// TIA Portal project "Log Control" (V20)

(* hardware
DEVICE "S7-1500/ET200MP station_1"  S7-1500 station
   slot 0: "Rail_0"  Rack  6ES7 590-1***0-0AA0
   slot 1: "PLC_1"  CPU 1518T-3 PN  6ES7 518-3TT10-0AB0  V4.0
      slot 3: "CPU display_1"  6ES7591-1BA00-0AA0
      slot 32768: "PROFINET interface_1"  X1
         slot 32769: "Port_1"  X1 P1
         slot 32770: "Port_2"  X1 P2
      slot 33024: "PROFINET interface_2"  X2
         slot 33025: "Port_1"  X2 P1
         slot 33026: "Port_2"  X2 P2
      slot 33280: "PROFINET interface GBIT_3"  X3
         slot 33281: "Port_1"  X3 P1
      slot 34817: "Virtual CP interface port_1"  Virtual CP interface port  Virtual CP interface port FW V4.0
DEVICE "LogHMI"  KTP700 Basic PN
   slot 0: "anit-hmi"  KTP700 Basic PN  6AV2 123-2GB03-0AX0  17.0.0.0
   slot 1: "HMI_RT_1"  KTP700 Basic PN  6AV2 123-2GB03-0AX0  17.0.0.0
   slot 5: "anit-hmi.IE_CP_1"  PROFINET Interface  17.0.0.0
      slot 1: "PROFINET Interface_1"  PROFINET Interface
         slot 1: "Port_1"  Port
*)

// ===== PLC "PLC_1"  CPU 1518T-3 PN =====
// protected blocks, not shown: "Log Control FC"

VAR_GLOBAL   // PLC tag table "Default tag table"
   "Tag_1" AT %M45.0 : Bool;
   "Tag_2" AT %M0.0 : Bool;
   "Tag_3" AT %M0.1 : Bool;
   "Tag_4" AT %M47.0 : Bool;
   "Tag_5" AT %M31.0 : Bool;
END_VAR

TYPE "LogControlUDT"
   STRUCT
      Settings : Struct
         "In Min" : Int := 0;
         "In Max" : Int := 100;
         "Out Min" : Real := 0.0;
         "Out Max" : Real := 100.0;
         "Log Repeat time" : Time := T#1s;
      END_STRUCT;
      "Worning Control" : Array[1..10] of Struct
         Text : String[20];
         MinValue : Real;
         MaxValue : Real;
      END_STRUCT;
      "Prescription Control" : Struct
         "Aktif Reçete" : Struct
            "Tarih/Saat" : DTL;
            Value : Real;
            Text : String;
         END_STRUCT;
         "Reçete Göstege" : Struct
            No : Array[0..10] of Int;
            "Tarih/Saat" : Array[0..10] of DTL;
            Value : Array[0..10] of Real;
            Text : Array[0..10] of String;
         END_STRUCT;
         T_ADD_Out : DTL;
         RET_Val_Out : DTL;
         p : Bool;
         "OP No" : Int;
         "OP Artı" : Bool;
         "OP Eksi" : Bool;
         "Gösterge No" : Int;
         "Gösterge Artı" : Bool;
         "Gösterge Eksi" : Bool;
         Log_Wride : Bool;
      END_STRUCT;
      Prescription : Array[0..101] of Struct
         "Tarih/Saat" : DTL;
         Value : Real;
         Text : String;
      END_STRUCT;
   END_STRUCT;
   // "Worning Control"[1].MinValue := 0.0;
   // "Worning Control"[1].MaxValue := 10.0;
   // "Worning Control"[1].Text := 'Value1';
   // "Worning Control"[2].Text := 'Value2';
   // "Worning Control"[2].MinValue := 10.0;
   // "Worning Control"[2].MaxValue := 20.0;
   // "Worning Control"[3].Text := 'Value3';
   // "Worning Control"[3].MinValue := 20.0;
   // "Worning Control"[3].MaxValue := 30.0;
   // "Worning Control"[4].Text := 'Value4';
   // "Worning Control"[4].MinValue := 30.0;
   // "Worning Control"[4].MaxValue := 40.0;
   // "Worning Control"[5].Text := 'Value5';
   // "Worning Control"[5].MinValue := 40.0;
   // "Worning Control"[5].MaxValue := 50.0;
   // "Worning Control"[6].Text := 'Value6';
   // "Worning Control"[6].MinValue := 50.0;
   // "Worning Control"[6].MaxValue := 60.0;
   // "Worning Control"[7].Text := 'Value7';
   // "Worning Control"[7].MinValue := 60.0;
   // "Worning Control"[7].MaxValue := 70.0;
   // "Worning Control"[8].Text := 'Value8';
   // "Worning Control"[8].MinValue := 70.0;
   // "Worning Control"[8].MaxValue := 80.0;
   // "Worning Control"[9].Text := 'Value9';
   // "Worning Control"[9].MinValue := 80.0;
   // "Worning Control"[9].MaxValue := 90.0;
   // "Worning Control"[10].Text := 'Value10';
   // "Worning Control"[10].MinValue := 90.0;
   // "Worning Control"[10].MaxValue := 100.0;
END_TYPE

DATA_BLOCK "Log Control DB"   // DB1
{ S7_Optimized_Access := 'TRUE' }
VERSION : 0.1
   VAR
      LogData : "LogControlUDT";
   END_VAR
BEGIN
END_DATA_BLOCK

// folder: 99-FuncLibrary

DATA_BLOCK "Value_1"   // DB4
{ S7_Optimized_Access := 'TRUE' }
VERSION : 0.1
   VAR
      InValue : Int;
      OutValue : Int;
      OutTime : DTL;
      OutText : String;
   END_VAR
BEGIN
END_DATA_BLOCK

// folder: System blocks/Program resources

DATA_BLOCK "IEC_Timer_0_DB"   // DB2
{ S7_Optimized_Access := 'TRUE' }
AUTHOR : Simatic
FAMILY : IEC
NAME : IEC_TMR
VERSION : 1.0
// stored: InstanceOfName IEC_TIMER
"IEC_TIMER"
BEGIN
END_DATA_BLOCK

DATA_BLOCK "IEC_Counter_0_DB"   // DB3
{ S7_Optimized_Access := 'TRUE' }
AUTHOR : Simatic
FAMILY : IEC
NAME : CNTR
VERSION : 1.0
// stored: InstanceOfName IEC_COUNTER
"IEC_COUNTER"
BEGIN
END_DATA_BLOCK

DATA_BLOCK "Value"   // DB5
{ S7_Optimized_Access := 'TRUE' }
AUTHOR : Simatic
FAMILY : IEC
NAME : IEC_TMR
VERSION : 1.0
// stored: InstanceOfName IEC_TIMER
"IEC_TIMER"
BEGIN
END_DATA_BLOCK

// folder: (top level)

ORGANIZATION_BLOCK "Main"   // OB1, LAD, ProgramCycle
TITLE = "Main Program Sweep (Cycle)"
{ S7_Optimized_Access := 'TRUE' }
VERSION : 0.1
   VAR_INPUT
      Initial_Call : Bool;   // Initial call of this OB
      Remanence : Bool;   // =True, if remanent data are available
   END_VAR
   VAR_TEMP
      Reset : Bool;
   END_VAR
   VAR_TEMP   // added for the SCL form of the ladder/FBD networks
      _w1 : Bool;
   END_VAR
BEGIN

REGION Network 1
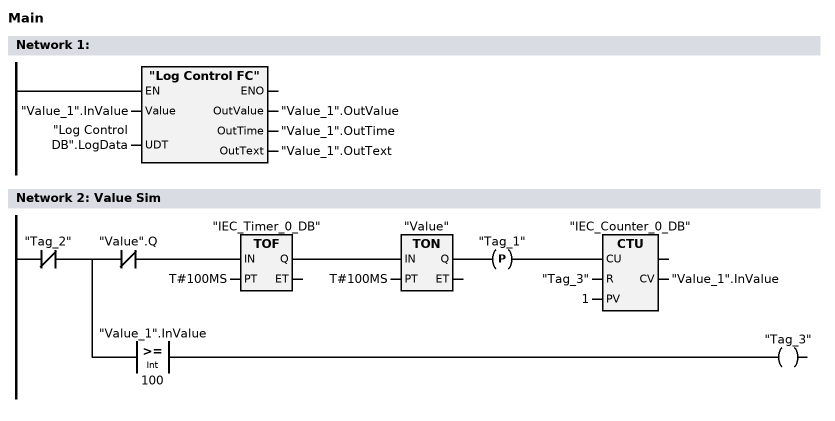
   RUNG wire#powerrail
      "Log Control FC"(Value := "Value_1".InValue, UDT := "Log Control DB".LogData, OutValue => "Value_1".OutValue, OutTime => "Value_1".OutTime, OutText => "Value_1".OutText)
   END_RUNG
   // the same network as SCL:
   "Log Control FC"(Value := "Value_1".InValue,
                    UDT := "Log Control DB".LogData,
                    OutValue => "Value_1".OutValue,
                    OutTime => "Value_1".OutTime,
                    OutText => "Value_1".OutText);
END_REGION

REGION Network 2: Value Sim
   "IEC_Timer_0_DB".TOF(IN := NOT "Tag_2" AND NOT "Value".Q, PT := T#100MS);
   "Value".TON(IN := "IEC_Timer_0_DB".Q, PT := T#100MS);
   #_w1 := "Value".Q AND NOT "Tag_1";   // rising edge
   "Tag_1" := "Value".Q;
   "IEC_Counter_0_DB".CTU(CU := #_w1, R := "Tag_3", PV := 1, CV => "Value_1".InValue);
   "Tag_3" := NOT "Tag_2" AND ("Value_1".InValue >= 100);
END_REGION
END_ORGANIZATION_BLOCK

(* ===== HMI "HMI_RT_1" =====
system functions are stored by id; their names below are inferred from use
connection "HMI_Connection_1": ETHERNET, SMART_S7_1500_OMS

HMI tags "Default tag table"
   "Log Control DB_LogData_Prescription Control_Reçete Göstege_No{1}" : Int = PLC "Log Control DB".LogData."Prescription Control"."Reçete Göstege".No[1], 100 ms
   "Log Control DB_LogData_Prescription Control_Reçete Göstege_No{2}" : Int = PLC "Log Control DB".LogData."Prescription Control"."Reçete Göstege".No[2], 100 ms
   "Log Control DB_LogData_Prescription Control_Reçete Göstege_No{3}" : Int = PLC "Log Control DB".LogData."Prescription Control"."Reçete Göstege".No[3], 100 ms
   "Log Control DB_LogData_Prescription Control_Reçete Göstege_No{4}" : Int = PLC "Log Control DB".LogData."Prescription Control"."Reçete Göstege".No[4], 100 ms
   "Log Control DB_LogData_Prescription Control_Reçete Göstege_No{5}" : Int = PLC "Log Control DB".LogData."Prescription Control"."Reçete Göstege".No[5], 100 ms
   "Log Control DB_LogData_Prescription Control_Reçete Göstege_No{6}" : Int = PLC "Log Control DB".LogData."Prescription Control"."Reçete Göstege".No[6], 100 ms
   "Log Control DB_LogData_Prescription Control_Reçete Göstege_No{7}" : Int = PLC "Log Control DB".LogData."Prescription Control"."Reçete Göstege".No[7], 100 ms
   "Log Control DB_LogData_Prescription Control_Reçete Göstege_No{8}" : Int = PLC "Log Control DB".LogData."Prescription Control"."Reçete Göstege".No[8], 100 ms
   "Log Control DB_LogData_Prescription Control_Reçete Göstege_No{9}" : Int = PLC "Log Control DB".LogData."Prescription Control"."Reçete Göstege".No[9], 100 ms
   "Log Control DB_LogData_Prescription Control_Reçete Göstege_No{10}" : Int = PLC "Log Control DB".LogData."Prescription Control"."Reçete Göstege".No[10], 100 ms
   "Log Control DB_LogData_Prescription Control_Reçete Göstege_Tarih/Saat{1}" : DTL = PLC "Log Control DB".LogData."Prescription Control"."Reçete Göstege".Tarih/Saat[1], 100 ms
   "Log Control DB_LogData_Prescription Control_Reçete Göstege_Tarih/Saat{2}" : DTL = PLC "Log Control DB".LogData."Prescription Control"."Reçete Göstege".Tarih/Saat[2], 100 ms
   "Log Control DB_LogData_Prescription Control_Reçete Göstege_Tarih/Saat{3}" : DTL = PLC "Log Control DB".LogData."Prescription Control"."Reçete Göstege".Tarih/Saat[3], 100 ms
   "Log Control DB_LogData_Prescription Control_Reçete Göstege_Tarih/Saat{4}" : DTL = PLC "Log Control DB".LogData."Prescription Control"."Reçete Göstege".Tarih/Saat[4], 100 ms
   "Log Control DB_LogData_Prescription Control_Reçete Göstege_Tarih/Saat{5}" : DTL = PLC "Log Control DB".LogData."Prescription Control"."Reçete Göstege".Tarih/Saat[5], 100 ms
   "Log Control DB_LogData_Prescription Control_Reçete Göstege_Tarih/Saat{6}" : DTL = PLC "Log Control DB".LogData."Prescription Control"."Reçete Göstege".Tarih/Saat[6], 100 ms
   "Log Control DB_LogData_Prescription Control_Reçete Göstege_Tarih/Saat{7}" : DTL = PLC "Log Control DB".LogData."Prescription Control"."Reçete Göstege".Tarih/Saat[7], 100 ms
   "Log Control DB_LogData_Prescription Control_Reçete Göstege_Tarih/Saat{8}" : DTL = PLC "Log Control DB".LogData."Prescription Control"."Reçete Göstege".Tarih/Saat[8], 100 ms
   "Log Control DB_LogData_Prescription Control_Reçete Göstege_Tarih/Saat{9}" : DTL = PLC "Log Control DB".LogData."Prescription Control"."Reçete Göstege".Tarih/Saat[9], 100 ms
   "Log Control DB_LogData_Prescription Control_Reçete Göstege_Tarih/Saat{10}" : DTL = PLC "Log Control DB".LogData."Prescription Control"."Reçete Göstege".Tarih/Saat[10], 100 ms
   "Log Control DB_LogData_Prescription Control_Reçete Göstege_Value{1}" : Real = PLC "Log Control DB".LogData."Prescription Control"."Reçete Göstege".Value[1], 100 ms
   "Log Control DB_LogData_Prescription Control_Reçete Göstege_Value{2}" : Real = PLC "Log Control DB".LogData."Prescription Control"."Reçete Göstege".Value[2], 100 ms
   "Log Control DB_LogData_Prescription Control_Reçete Göstege_Value{3}" : Real = PLC "Log Control DB".LogData."Prescription Control"."Reçete Göstege".Value[3], 100 ms
   "Log Control DB_LogData_Prescription Control_Reçete Göstege_Value{4}" : Real = PLC "Log Control DB".LogData."Prescription Control"."Reçete Göstege".Value[4], 100 ms
   "Log Control DB_LogData_Prescription Control_Reçete Göstege_Value{5}" : Real = PLC "Log Control DB".LogData."Prescription Control"."Reçete Göstege".Value[5], 100 ms
   "Log Control DB_LogData_Prescription Control_Reçete Göstege_Value{6}" : Real = PLC "Log Control DB".LogData."Prescription Control"."Reçete Göstege".Value[6], 100 ms
   "Log Control DB_LogData_Prescription Control_Reçete Göstege_Value{7}" : Real = PLC "Log Control DB".LogData."Prescription Control"."Reçete Göstege".Value[7], 100 ms
   "Log Control DB_LogData_Prescription Control_Reçete Göstege_Value{8}" : Real = PLC "Log Control DB".LogData."Prescription Control"."Reçete Göstege".Value[8], 100 ms
   "Log Control DB_LogData_Prescription Control_Reçete Göstege_Value{9}" : Real = PLC "Log Control DB".LogData."Prescription Control"."Reçete Göstege".Value[9], 100 ms
   "Log Control DB_LogData_Prescription Control_Reçete Göstege_Value{10}" : Real = PLC "Log Control DB".LogData."Prescription Control"."Reçete Göstege".Value[10], 100 ms
   "Log Control DB_LogData_Prescription Control_Reçete Göstege_Text{1}" : String[254] = PLC "Log Control DB".LogData."Prescription Control"."Reçete Göstege".Text[1], 100 ms
   "Log Control DB_LogData_Prescription Control_Reçete Göstege_Text{2}" : String[254] = PLC "Log Control DB".LogData."Prescription Control"."Reçete Göstege".Text[2], 100 ms
   "Log Control DB_LogData_Prescription Control_Reçete Göstege_Text{3}" : String[254] = PLC "Log Control DB".LogData."Prescription Control"."Reçete Göstege".Text[3], 100 ms
   "Log Control DB_LogData_Prescription Control_Reçete Göstege_Text{4}" : String[254] = PLC "Log Control DB".LogData."Prescription Control"."Reçete Göstege".Text[4], 100 ms
   "Log Control DB_LogData_Prescription Control_Reçete Göstege_Text{5}" : String[254] = PLC "Log Control DB".LogData."Prescription Control"."Reçete Göstege".Text[5], 100 ms
   "Log Control DB_LogData_Prescription Control_Reçete Göstege_Text{6}" : String[254] = PLC "Log Control DB".LogData."Prescription Control"."Reçete Göstege".Text[6], 100 ms
   "Log Control DB_LogData_Prescription Control_Reçete Göstege_Text{7}" : String[254] = PLC "Log Control DB".LogData."Prescription Control"."Reçete Göstege".Text[7], 100 ms
   "Log Control DB_LogData_Prescription Control_Reçete Göstege_Text{8}" : String[254] = PLC "Log Control DB".LogData."Prescription Control"."Reçete Göstege".Text[8], 100 ms
   "Log Control DB_LogData_Prescription Control_Reçete Göstege_Text{9}" : String[254] = PLC "Log Control DB".LogData."Prescription Control"."Reçete Göstege".Text[9], 100 ms
   "Log Control DB_LogData_Prescription Control_Reçete Göstege_Text{10}" : String[254] = PLC "Log Control DB".LogData."Prescription Control"."Reçete Göstege".Text[10], 100 ms
   "Log Control DB_LogData_Prescription Control_Gösterge Artı" : Bool = PLC "Log Control DB".LogData."Prescription Control"."Gösterge Artı", 100 ms
   "Log Control DB_LogData_Prescription Control_Gösterge Eksi" : Bool = PLC "Log Control DB".LogData."Prescription Control"."Gösterge Eksi", 100 ms

discrete alarms
   1: 'Acil Stop Basılı', class I-Shaft, trigger "Alarm_A1{0}" bit 0
   2: 'Shaft Kilit İleri Gidemedi', class I-Shaft, trigger "Alarm_A1{0}" bit 1
   3: 'Shaft Kilit Geri Gidemedi', class I-Shaft, trigger "Alarm_A1{0}" bit 2
   4: 'Gövde Kilit İleri Gidemedi', class I-Shaft, trigger "Alarm_A1{0}" bit 3
   5: 'Gövde Kilit Geri Gidemedi', class I-Shaft, trigger "Alarm_A1{0}" bit 4
   6: 'Shaft Kamera TimeOut', class I-Shaft, trigger "Alarm_A1{0}" bit 5
   7: 'Civata Kamera TimeOut', class I-Shaft, trigger "Alarm_A1{0}" bit 6
   8: 'Shaft Kamera Hata', class I-Shaft, trigger "Alarm_A1{0}" bit 7
   9: 'Civata Kamera Hata', class I-Shaft, trigger "Alarm_A1{0}" bit 8
   10: '-', class I-Shaft, trigger "Alarm_A1{0}" bit 9
   11: '-', class I-Shaft, trigger "Alarm_A1{0}" bit 10
   12: '-', class I-Shaft, trigger "Alarm_A1{0}" bit 11
   13: '-', class I-Shaft, trigger "Alarm_A1{0}" bit 12
   14: '-', class I-Shaft, trigger "Alarm_A1{0}" bit 13
   15: '-', class I-Shaft, trigger "Alarm_A1{0}" bit 14
   16: '-', class I-Shaft, trigger "Alarm_A1{0}" bit 15
   17: 'Konveyör Yükleme Bölgesi Acil Stop Basılı', class Konveyör, trigger "Alarm_A1{1}" bit 0
   18: 'Konveyör Çıkış Bölgesi Acil Stop Basılı', class Konveyör, trigger "Alarm_A1{1}" bit 1
   19: 'Ürün İstenen Konumdan Çok İleri Gitti.Ürünü Alıp Reset Butonuna Basınız.İlgili Sensörü Kontrol Ediniz.', class Konveyör, trigger "Alarm_A1{1}" bit 2
   20: 'Konveyör İstasyon 3 Ürün Düzgün Oturmadı Hatası, Ürünü Düzeltiniz, Konveyör Sayfasından Hatayı Resetleyiniz', class Konveyör, trigger "Alarm_A1{1}" bit 3
   21: 'Konveyör İstasyon 4 Ürün Düzgün Oturmadı Hatası, Ürünü Düzeltiniz, Konveyör Sayfasından Hatayı Resetleyiniz', class Konveyör, trigger "Alarm_A1{1}" bit 4
   22: 'Konveyör İstasyon 5 Ürün Düzgün Oturmadı Hatası, Ürünü Düzeltiniz, Konveyör Sayfasından Hatayı Resetleyiniz', class Konveyör, trigger "Alarm_A1{1}" bit 5
   23: 'Konveyör İstasyon 6 Ürün Düzgün Oturmadı Hatası, Ürünü Düzeltiniz, Konveyör Sayfasından Hatayı Resetleyiniz', class Konveyör, trigger "Alarm_A1{1}" bit 6
   24: 'Konveyör İstasyon 1 Ürün Düzgün Oturmadı Hatası, Ürünü Düzeltiniz, Konveyör Sayfasından Hatayı Resetleyiniz', class Konveyör, trigger "Alarm_A1{1}" bit 7

screen "01 - Company" 800x480, template "Main Template_Anasayfa"
   TextField "Text field_1" at 28,18 size 61x23; Text 'Log No / Kayıt No:'
   IOField "I/O field_1" at 29,53 size 65x33; FormatPattern 999
      ProcessValue <- "Log Control DB_LogData_Prescription Control_Reçete Göstege_No{1}"
   Button "Button_1" at 497,417 size 142x57; TextOff '<< / >>'
      on Press: function_b14e0dd5("Log Control DB_LogData_Prescription Control_Gösterge Eksi", 0)
   Button "Button_2" at 653,417 size 142x57; TextOff '>> / <<'
      on Press: function_b14e0dd5("Log Control DB_LogData_Prescription Control_Gösterge Artı", 0)
   IOField "I/O field_2" at 29,88 size 65x33; FormatPattern 999
      ProcessValue <- "Log Control DB_LogData_Prescription Control_Reçete Göstege_No{2}"
   IOField "I/O field_5" at 29,123 size 65x33; FormatPattern 999
      ProcessValue <- "Log Control DB_LogData_Prescription Control_Reçete Göstege_No{3}"
   IOField "I/O field_7" at 29,158 size 65x33; FormatPattern 999
      ProcessValue <- "Log Control DB_LogData_Prescription Control_Reçete Göstege_No{4}"
   IOField "I/O field_9" at 29,193 size 65x33; FormatPattern 999
      ProcessValue <- "Log Control DB_LogData_Prescription Control_Reçete Göstege_No{5}"
   IOField "I/O field_11" at 29,229 size 65x33; FormatPattern 999
      ProcessValue <- "Log Control DB_LogData_Prescription Control_Reçete Göstege_No{6}"
   IOField "I/O field_13" at 29,264 size 65x33; FormatPattern 999
      ProcessValue <- "Log Control DB_LogData_Prescription Control_Reçete Göstege_No{7}"
   IOField "I/O field_15" at 29,299 size 65x33; FormatPattern 999
      ProcessValue <- "Log Control DB_LogData_Prescription Control_Reçete Göstege_No{8}"
   IOField "I/O field_17" at 29,334 size 65x33; FormatPattern 999
      ProcessValue <- "Log Control DB_LogData_Prescription Control_Reçete Göstege_No{9}"
   IOField "I/O field_19" at 29,370 size 65x33; FormatPattern 999
      ProcessValue <- "Log Control DB_LogData_Prescription Control_Reçete Göstege_No{10}"
   IOField "I/O field_26" at 108,54 size 183x32; FormatPattern 9999999999999999999999999999999999999999
      ProcessValue <- "Log Control DB_LogData_Prescription Control_Reçete Göstege_Tarih/Saat{1}"
   IOField "I/O field_3" at 108,89 size 183x32; FormatPattern 9999999999999999999999999999999999999999
      ProcessValue <- "Log Control DB_LogData_Prescription Control_Reçete Göstege_Tarih/Saat{2}"
   IOField "I/O field_4" at 108,124 size 183x32; FormatPattern 9999999999999999999999999999999999999999
      ProcessValue <- "Log Control DB_LogData_Prescription Control_Reçete Göstege_Tarih/Saat{3}"
   IOField "I/O field_6" at 108,159 size 183x32; FormatPattern 9999999999999999999999999999999999999999
      ProcessValue <- "Log Control DB_LogData_Prescription Control_Reçete Göstege_Tarih/Saat{4}"
   IOField "I/O field_8" at 108,194 size 183x32; FormatPattern 9999999999999999999999999999999999999999
      ProcessValue <- "Log Control DB_LogData_Prescription Control_Reçete Göstege_Tarih/Saat{5}"
   IOField "I/O field_10" at 108,230 size 183x32; FormatPattern 9999999999999999999999999999999999999999
      ProcessValue <- "Log Control DB_LogData_Prescription Control_Reçete Göstege_Tarih/Saat{6}"
   IOField "I/O field_12" at 108,265 size 183x32; FormatPattern 9999999999999999999999999999999999999999
      ProcessValue <- "Log Control DB_LogData_Prescription Control_Reçete Göstege_Tarih/Saat{7}"
   IOField "I/O field_14" at 108,300 size 183x32; FormatPattern 9999999999999999999999999999999999999999
      ProcessValue <- "Log Control DB_LogData_Prescription Control_Reçete Göstege_Tarih/Saat{8}"
   IOField "I/O field_16" at 108,335 size 183x32; FormatPattern 9999999999999999999999999999999999999999
      ProcessValue <- "Log Control DB_LogData_Prescription Control_Reçete Göstege_Tarih/Saat{9}"
   IOField "I/O field_18" at 108,371 size 183x32; FormatPattern 9999999999999999999999999999999999999999
      ProcessValue <- "Log Control DB_LogData_Prescription Control_Reçete Göstege_Tarih/Saat{10}"
   TextField "Text field_2" at 160,18 size 80x23; Text 'Log Time / Kayıt No:'
   TextField "Text field_3" at 339,18 size 85x23; Text 'Log Value / Kayıt No:'
   IOField "I/O field_20" at 302,53 size 159x33; FormatPattern 9999.999
      ProcessValue <- "Log Control DB_LogData_Prescription Control_Reçete Göstege_Value{1}"
   TextField "Text field_4" at 596,18 size 77x23; Text 'Log Text / Kayıt No:'
   IOField "I/O field_21" at 480,53 size 308x33; FormatPattern ????????????????????
      ProcessValue <- "Log Control DB_LogData_Prescription Control_Reçete Göstege_Text{1}"
   IOField "I/O field_22" at 302,88 size 159x33; FormatPattern 9999.999
      ProcessValue <- "Log Control DB_LogData_Prescription Control_Reçete Göstege_Value{2}"
   IOField "I/O field_23" at 480,88 size 308x33; FormatPattern ????????????????????
      ProcessValue <- "Log Control DB_LogData_Prescription Control_Reçete Göstege_Text{2}"
   IOField "I/O field_24" at 302,123 size 159x33; FormatPattern 9999.999
      ProcessValue <- "Log Control DB_LogData_Prescription Control_Reçete Göstege_Value{3}"
   IOField "I/O field_25" at 480,123 size 308x33; FormatPattern ????????????????????
      ProcessValue <- "Log Control DB_LogData_Prescription Control_Reçete Göstege_Text{3}"
   IOField "I/O field_27" at 302,158 size 159x33; FormatPattern 9999.999
      ProcessValue <- "Log Control DB_LogData_Prescription Control_Reçete Göstege_Value{4}"
   IOField "I/O field_28" at 480,158 size 308x33; FormatPattern ????????????????????
      ProcessValue <- "Log Control DB_LogData_Prescription Control_Reçete Göstege_Text{4}"
   IOField "I/O field_29" at 302,193 size 159x33; FormatPattern 9999.999
      ProcessValue <- "Log Control DB_LogData_Prescription Control_Reçete Göstege_Value{5}"
   IOField "I/O field_30" at 480,193 size 308x33; FormatPattern ????????????????????
      ProcessValue <- "Log Control DB_LogData_Prescription Control_Reçete Göstege_Text{5}"
   IOField "I/O field_31" at 302,229 size 159x33; FormatPattern 9999.999
      ProcessValue <- "Log Control DB_LogData_Prescription Control_Reçete Göstege_Value{6}"
   IOField "I/O field_32" at 480,229 size 308x33; FormatPattern ????????????????????
      ProcessValue <- "Log Control DB_LogData_Prescription Control_Reçete Göstege_Text{6}"
   IOField "I/O field_33" at 302,264 size 159x33; FormatPattern 9999.999
      ProcessValue <- "Log Control DB_LogData_Prescription Control_Reçete Göstege_Value{7}"
   IOField "I/O field_34" at 480,264 size 308x33; FormatPattern ????????????????????
      ProcessValue <- "Log Control DB_LogData_Prescription Control_Reçete Göstege_Text{7}"
   IOField "I/O field_35" at 302,299 size 159x33; FormatPattern 9999.999
      ProcessValue <- "Log Control DB_LogData_Prescription Control_Reçete Göstege_Value{8}"
   IOField "I/O field_36" at 480,299 size 308x33; FormatPattern ????????????????????
      ProcessValue <- "Log Control DB_LogData_Prescription Control_Reçete Göstege_Text{8}"
   IOField "I/O field_37" at 302,334 size 159x33; FormatPattern 9999.999
      ProcessValue <- "Log Control DB_LogData_Prescription Control_Reçete Göstege_Value{9}"
   IOField "I/O field_38" at 480,334 size 308x33; FormatPattern ????????????????????
      ProcessValue <- "Log Control DB_LogData_Prescription Control_Reçete Göstege_Text{9}"
   IOField "I/O field_39" at 302,370 size 159x33; FormatPattern 9999.999
      ProcessValue <- "Log Control DB_LogData_Prescription Control_Reçete Göstege_Value{10}"
   IOField "I/O field_40" at 480,370 size 308x33; FormatPattern ????????????????????
      ProcessValue <- "Log Control DB_LogData_Prescription Control_Reçete Göstege_Text{10}"

Template "Main Template" 800x480
   TextField "Template_Text field_1" at 0,460 size 100x20; Text 'Firma'
   TextField "Template_Text field_2" at 100,460 size 100x20; Text 'Anasayfa'
   TextField "Template_Text field_3" at 200,460 size 100x20; Text 'Manuel'
   TextField "Template_Text field_4" at 300,460 size 100x20; Text 'PLC Input'
   TextField "Template_Text field_5" at 400,460 size 100x20; Text 'PLC Output'
   TextField "Template_Text field_6" at 500,460 size 100x20; Text 'Ayarlar'
   TextField "Template_Text field_7" at 600,460 size 100x20; Text 'G. Alarmlar'
   TextField "Template_Text field_8" at 700,460 size 100x20; Text 'Alarmlar'
   GraphicView "Template_Graphic view_2" at 611,3 size 184x40; Picture "panel-makotim-logo-buyuk"
   DateTimeField "Template_Date/time field_2" at 570,43 size 225x23
*)